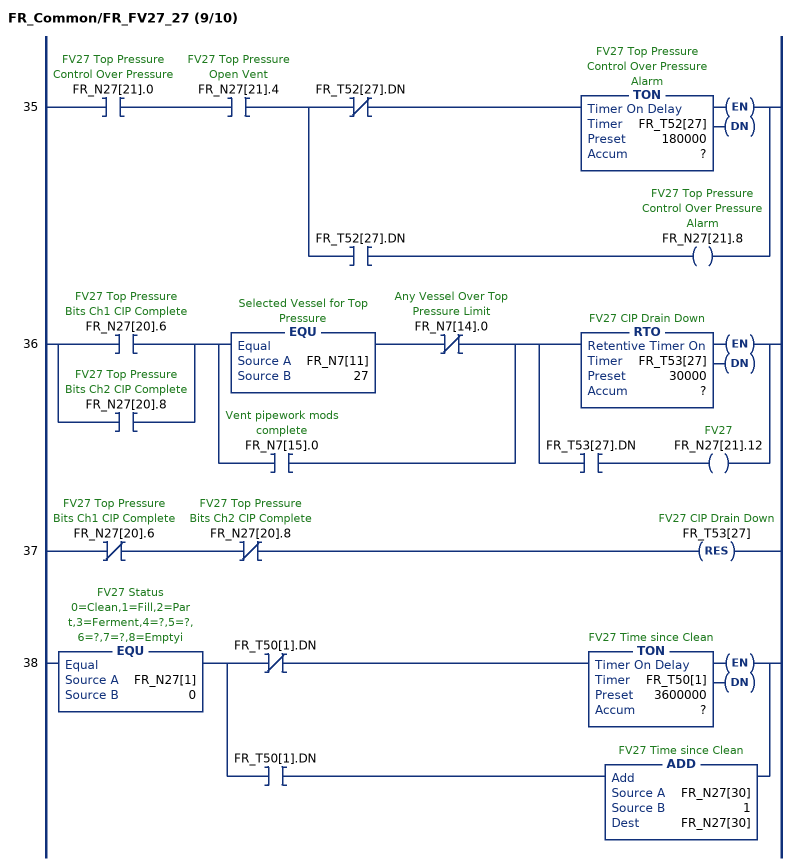
   35: XIC(FR_N27[21].0)XIC(FR_N27[21].4)[XIO(FR_T52[27].DN) TON(FR_T52[27],?,?) ,XIC(FR_T52[27].DN) OTE(FR_N27[21].8) ];
   36: [XIC(FR_N27[20].6) ,XIC(FR_N27[20].8) ][EQU(FR_N7[11],27) XIO(FR_N7[14].0) ,XIC(FR_N7[15].0) ][RTO(FR_T53[27],?,?) ,XIC(FR_T53[27].DN) OTE(FR_N27[21].12) ];
   37: XIO(FR_N27[20].6)XIO(FR_N27[20].8)RES(FR_T53[27]);
   38: EQU(FR_N27[1],0)[XIO(FR_T50[1].DN) TON(FR_T50[1],?,?) ,XIC(FR_T50[1].DN) ADD(FR_N27[30],1,FR_N27[30]) ];
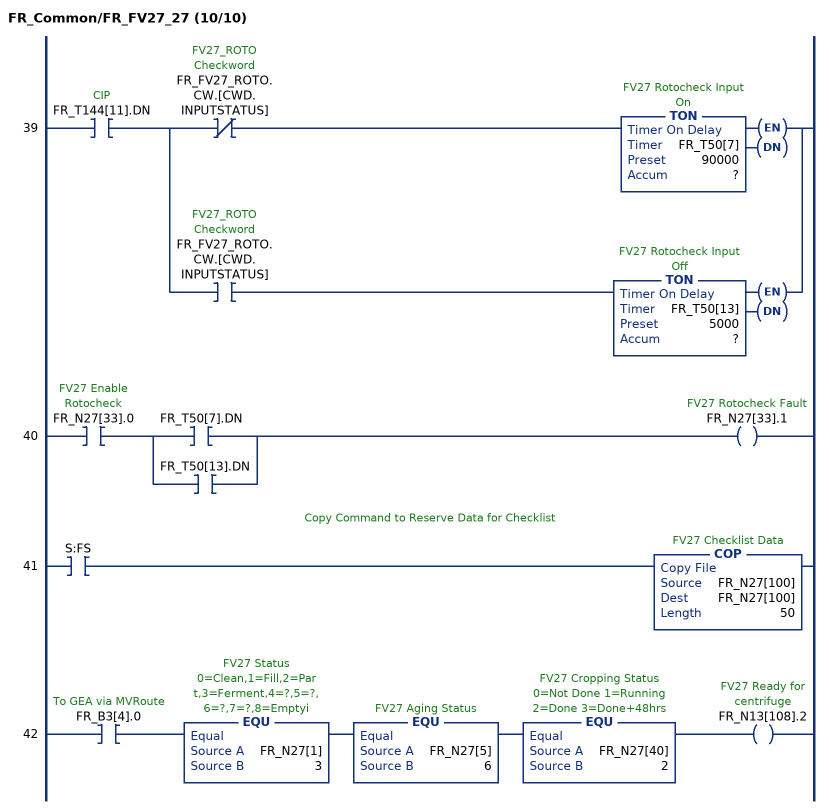
   39: XIC(FR_T144[11].DN)[XIO(FR_FV27_ROTO.CW.[CWD.INPUTSTATUS]) TON(FR_T50[7],?,?) ,XIC(FR_FV27_ROTO.CW.[CWD.INPUTSTATUS]) TON(FR_T50[13],?,?) ];
   40: XIC(FR_N27[33].0)[XIC(FR_T50[7].DN) ,XIC(FR_T50[13].DN) ]OTE(FR_N27[33].1);
   // Copy Command to Reserve Data for Checklist
   41: XIC(S:FS)COP(FR_N27[100],FR_N27[100],50);
   42: XIC(FR_B3[4].0)EQU(FR_N27[1],3)EQU(FR_N27[5],6)EQU(FR_N27[40],2)OTE(FR_N13[108].2);
END_ROUTINE

ROUTINE FR_FV28_28   (* ladder *)
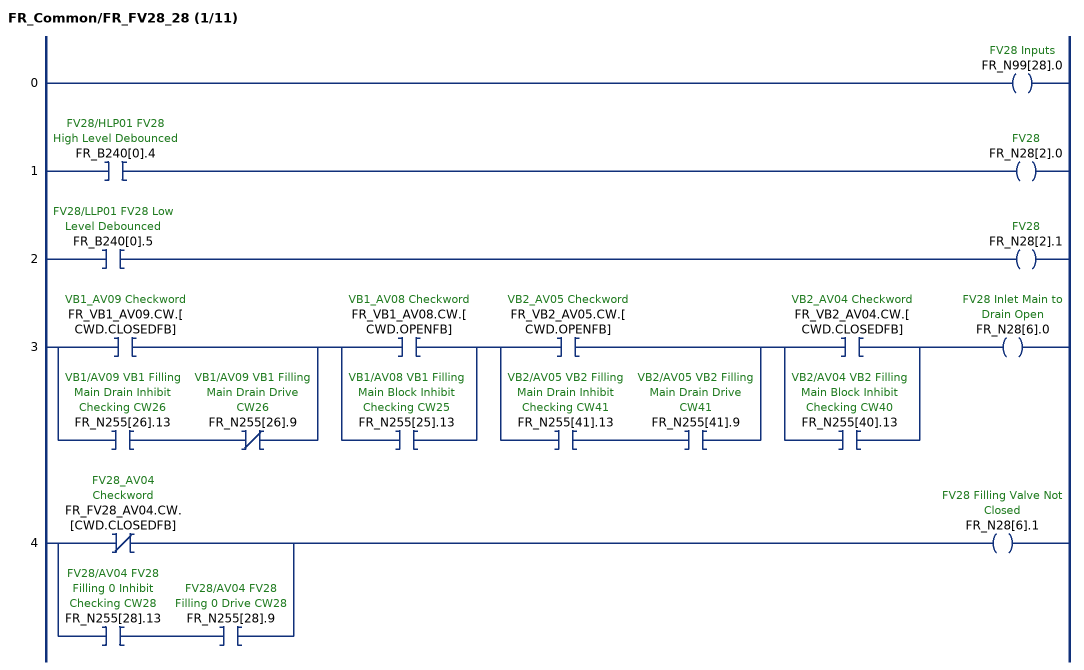
   0: OTE(FR_N99[28].0);
   1: XIC(FR_B240[0].4)OTE(FR_N28[2].0);
   2: XIC(FR_B240[0].5)OTE(FR_N28[2].1);
   3: [XIC(FR_VB1_AV09.CW.[CWD.CLOSEDFB]) ,XIC(FR_N255[26].13) XIO(FR_N255[26].9) ][XIC(FR_VB1_AV08.CW.[CWD.OPENFB]) ,XIC(FR_N255[25].13) ][XIC(FR_VB2_AV05.CW.[CWD.OPENFB]) ,XIC(FR_N255[41].13) XIC(FR_N255[41].9) ][XIC(FR_VB2_AV04.CW.[CWD.CLOSEDFB]) ,XIC(FR_N255[40].13) ]OTE(FR_N28[6].0);
   4: [XIO(FR_FV28_AV04.CW.[CWD.CLOSEDFB]) ,XIC(FR_N255[28].13) XIC(FR_N255[28].9) ]OTE(FR_N28[6].1);
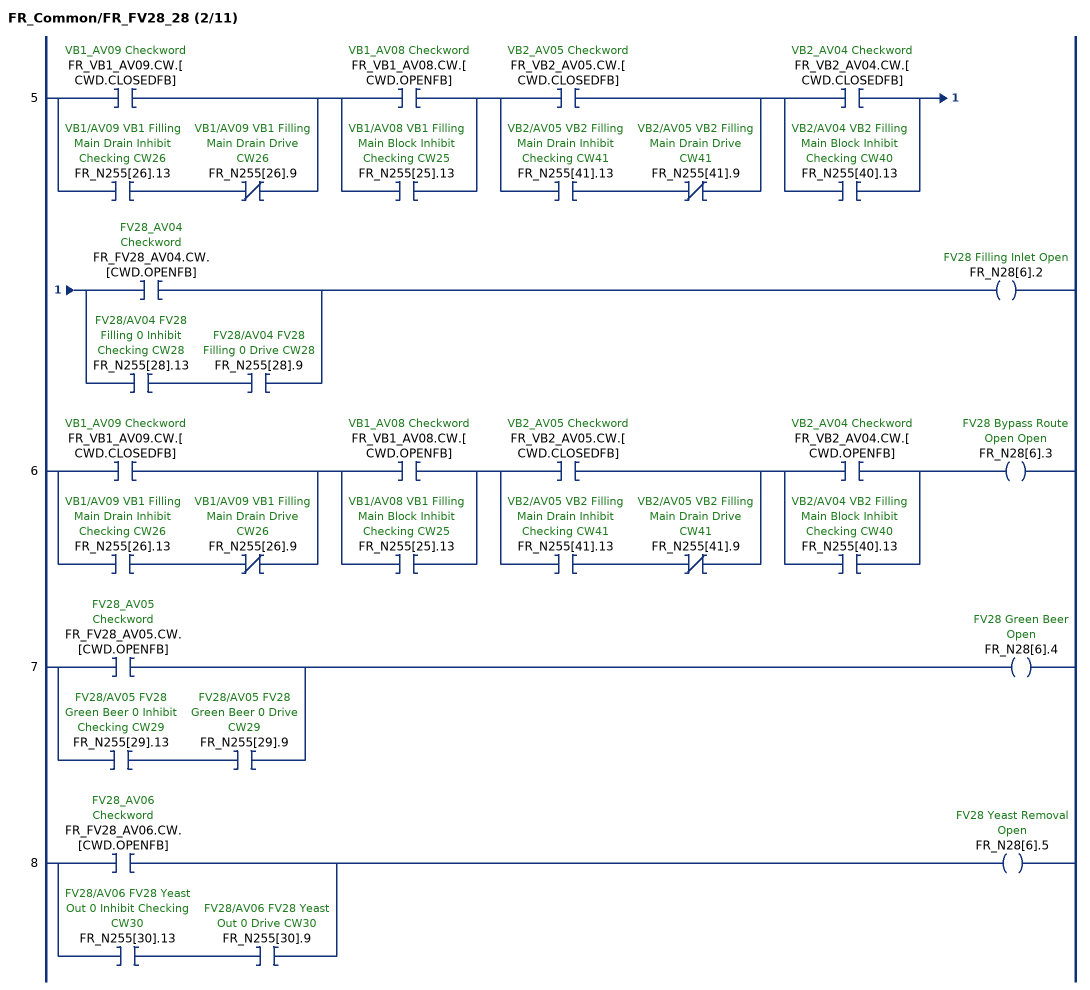
   5: [XIC(FR_VB1_AV09.CW.[CWD.CLOSEDFB]) ,XIC(FR_N255[26].13) XIO(FR_N255[26].9) ][XIC(FR_VB1_AV08.CW.[CWD.OPENFB]) ,XIC(FR_N255[25].13) ][XIC(FR_VB2_AV05.CW.[CWD.CLOSEDFB]) ,XIC(FR_N255[41].13) XIO(FR_N255[41].9) ][XIC(FR_VB2_AV04.CW.[CWD.CLOSEDFB]) ,XIC(FR_N255[40].13) ][XIC(FR_FV28_AV04.CW.[CWD.OPENFB]) ,XIC(FR_N255[28].13) XIC(FR_N255[28].9) ]OTE(FR_N28[6].2);
   6: [XIC(FR_VB1_AV09.CW.[CWD.CLOSEDFB]) ,XIC(FR_N255[26].13) XIO(FR_N255[26].9) ][XIC(FR_VB1_AV08.CW.[CWD.OPENFB]) ,XIC(FR_N255[25].13) ][XIC(FR_VB2_AV05.CW.[CWD.CLOSEDFB]) ,XIC(FR_N255[41].13) XIO(FR_N255[41].9) ][XIC(FR_VB2_AV04.CW.[CWD.OPENFB]) ,XIC(FR_N255[40].13) ]OTE(FR_N28[6].3);
   7: [XIC(FR_FV28_AV05.CW.[CWD.OPENFB]) ,XIC(FR_N255[29].13) XIC(FR_N255[29].9) ]OTE(FR_N28[6].4);
   8: [XIC(FR_FV28_AV06.CW.[CWD.OPENFB]) ,XIC(FR_N255[30].13) XIC(FR_N255[30].9) ]OTE(FR_N28[6].5);
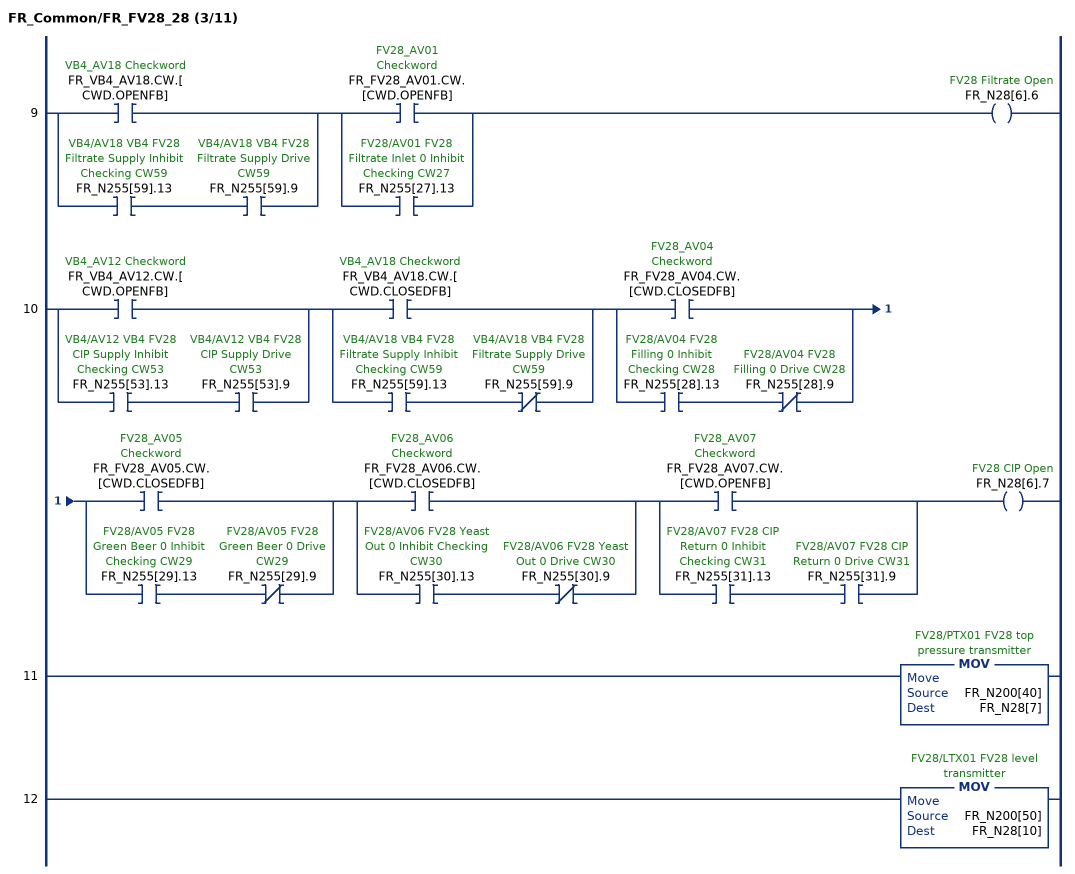
   9: [XIC(FR_VB4_AV18.CW.[CWD.OPENFB]) ,XIC(FR_N255[59].13) XIC(FR_N255[59].9) ][XIC(FR_FV28_AV01.CW.[CWD.OPENFB]) ,XIC(FR_N255[27].13) ]OTE(FR_N28[6].6);
   10: [XIC(FR_VB4_AV12.CW.[CWD.OPENFB]) ,XIC(FR_N255[53].13) XIC(FR_N255[53].9) ][XIC(FR_VB4_AV18.CW.[CWD.CLOSEDFB]) ,XIC(FR_N255[59].13) XIO(FR_N255[59].9) ][XIC(FR_FV28_AV04.CW.[CWD.CLOSEDFB]) ,XIC(FR_N255[28].13) XIO(FR_N255[28].9) ][XIC(FR_FV28_AV05.CW.[CWD.CLOSEDFB]) ,XIC(FR_N255[29].13) XIO(FR_N255[29].9) ][XIC(FR_FV28_AV06.CW.[CWD.CLOSEDFB]) ,XIC(FR_N255[30].13) XIO(FR_N255[30].9) ][XIC(FR_FV28_AV07.CW.[CWD.OPENFB]) ,XIC(FR_N255[31].13) XIC(FR_N255[31].9) ]OTE(FR_N28[6].7);
   11: MOV(FR_N200[40],FR_N28[7]);
   12: MOV(FR_N200[50],FR_N28[10]);
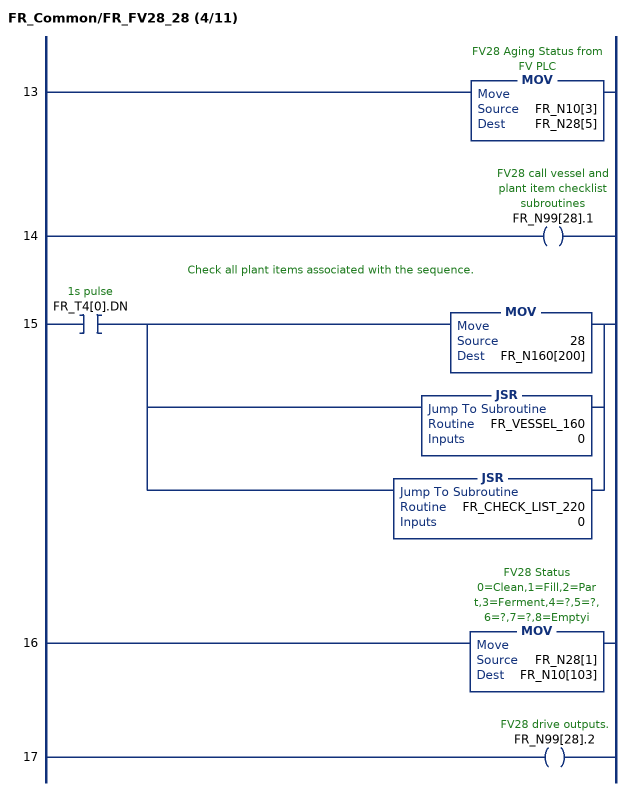
   13: MOV(FR_N10[3],FR_N28[5]);
   14: OTE(FR_N99[28].1);
   // Check all plant items associated with the sequence.
   15: XIC(FR_T4[0].DN)[MOV(28,FR_N160[200]) ,JSR(FR_VESSEL_160,0) ,JSR(FR_CHECK_LIST_220,0) ];
   16: MOV(FR_N28[1],FR_N10[103]);
   17: OTE(FR_N99[28].2);
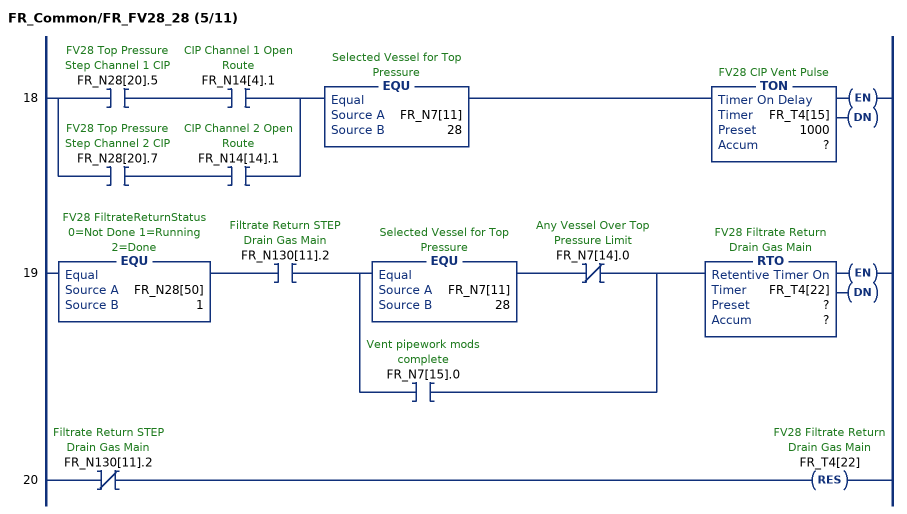
   18: [XIC(FR_N28[20].5) XIC(FR_N14[4].1) ,XIC(FR_N28[20].7) XIC(FR_N14[14].1) ]EQU(FR_N7[11],28)TON(FR_T4[15],?,?);
   19: EQU(FR_N28[50],1)XIC(FR_N130[11].2)[EQU(FR_N7[11],28) XIO(FR_N7[14].0) ,XIC(FR_N7[15].0) ]RTO(FR_T4[22],?,?);
   20: XIO(FR_N130[11].2)RES(FR_T4[22]);
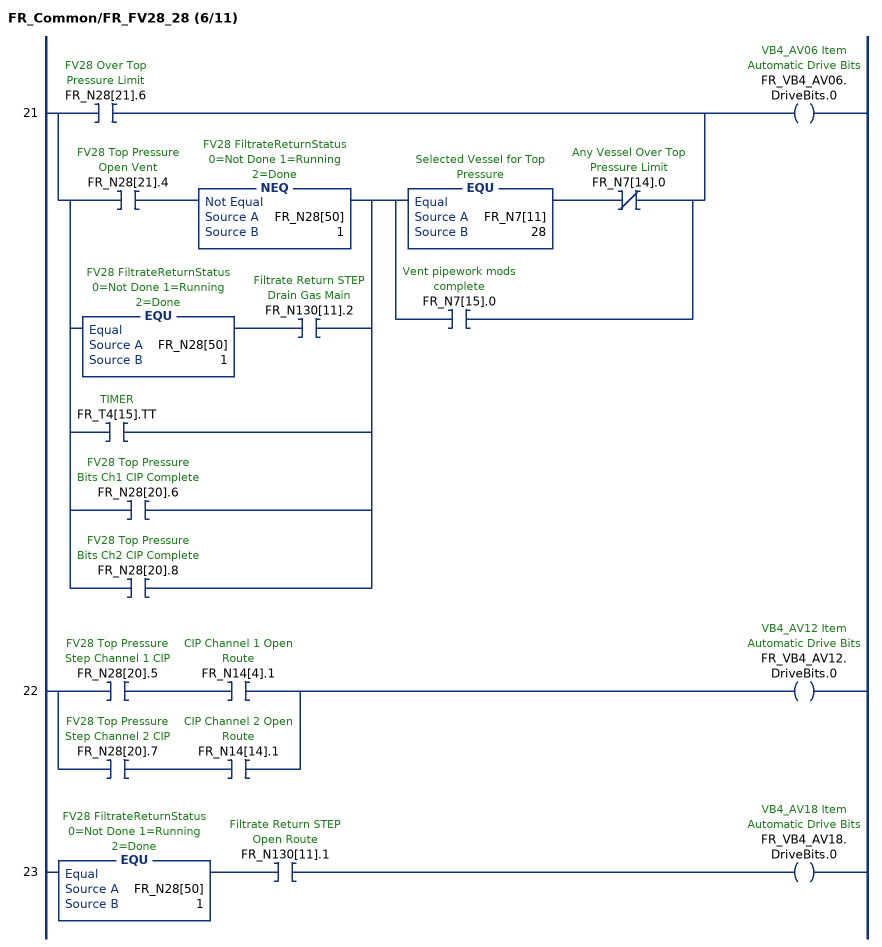
   21: [XIC(FR_N28[21].6) ,[XIC(FR_N28[21].4) NEQ(FR_N28[50],1) ,EQU(FR_N28[50],1) XIC(FR_N130[11].2) ,XIC(FR_T4[15].TT) ,[XIC(FR_N28[20].6) ,XIC(FR_N28[20].8) ] ] [EQU(FR_N7[11],28) XIO(FR_N7[14].0) ,XIC(FR_N7[15].0) ] ]OTE(FR_VB4_AV06.DriveBits.0);
   22: [XIC(FR_N28[20].5) XIC(FR_N14[4].1) ,XIC(FR_N28[20].7) XIC(FR_N14[14].1) ]OTE(FR_VB4_AV12.DriveBits.0);
   23: EQU(FR_N28[50],1)XIC(FR_N130[11].1)OTE(FR_VB4_AV18.DriveBits.0);
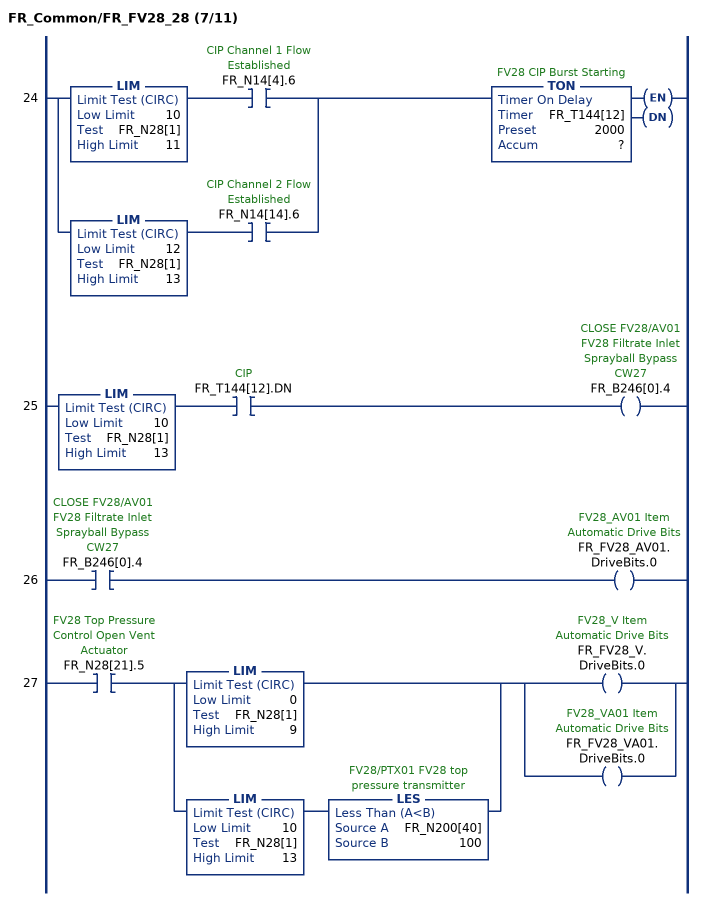
   24: [LIM(10,FR_N28[1],11) XIC(FR_N14[4].6) ,LIM(12,FR_N28[1],13) XIC(FR_N14[14].6) ]TON(FR_T144[12],?,?);
   25: LIM(10,FR_N28[1],13)XIC(FR_T144[12].DN)OTE(FR_B246[0].4);
   26: XIC(FR_B246[0].4)OTE(FR_FV28_AV01.DriveBits.0);
   27: XIC(FR_N28[21].5)[LIM(0,FR_N28[1],9) ,LIM(10,FR_N28[1],13) LES(FR_N200[40],100) ][OTE(FR_FV28_V.DriveBits.0) ,OTE(FR_FV28_VA01.DriveBits.0) ];
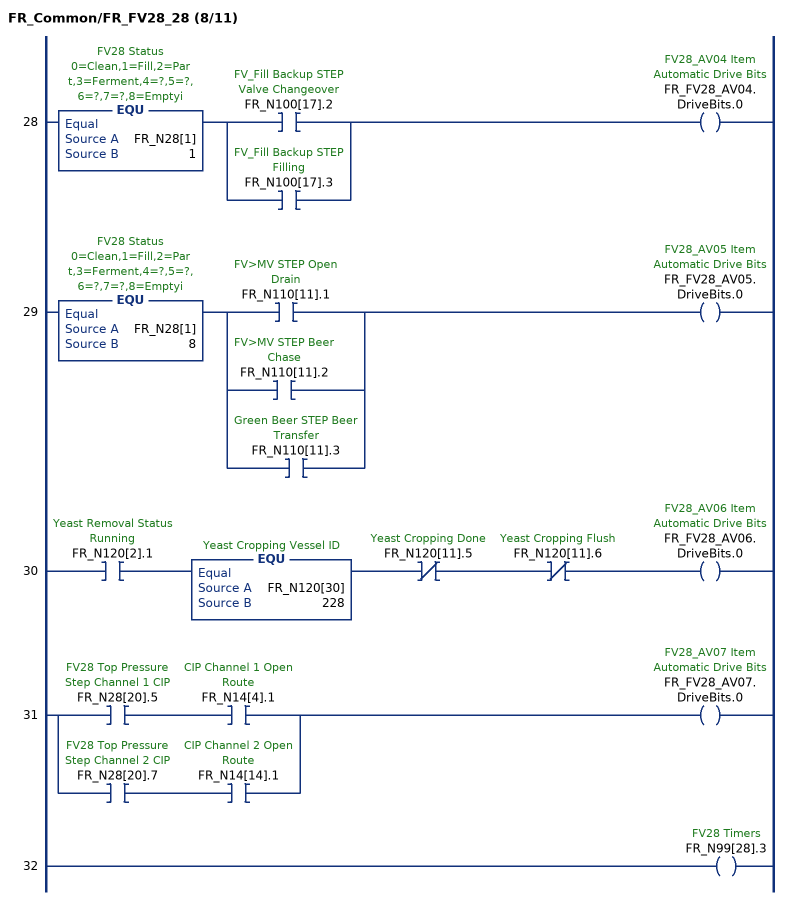
   28: EQU(FR_N28[1],1)[XIC(FR_N100[17].2) ,XIC(FR_N100[17].3) ]OTE(FR_FV28_AV04.DriveBits.0);
   29: EQU(FR_N28[1],8)[XIC(FR_N110[11].1) ,XIC(FR_N110[11].2) ,XIC(FR_N110[11].3) ]OTE(FR_FV28_AV05.DriveBits.0);
   30: XIC(FR_N120[2].1)EQU(FR_N120[30],228)XIO(FR_N120[11].5)XIO(FR_N120[11].6)OTE(FR_FV28_AV06.DriveBits.0);
   31: [XIC(FR_N28[20].5) XIC(FR_N14[4].1) ,XIC(FR_N28[20].7) XIC(FR_N14[14].1) ]OTE(FR_FV28_AV07.DriveBits.0);
   32: OTE(FR_N99[28].3);
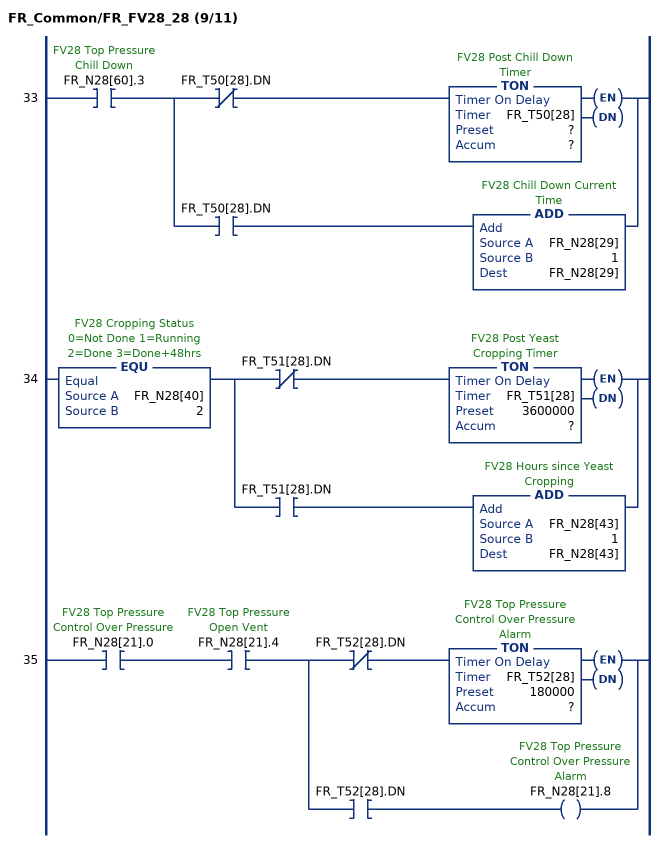
   33: XIC(FR_N28[60].3)[XIO(FR_T50[28].DN) TON(FR_T50[28],?,?) ,XIC(FR_T50[28].DN) ADD(FR_N28[29],1,FR_N28[29]) ];
   34: EQU(FR_N28[40],2)[XIO(FR_T51[28].DN) TON(FR_T51[28],?,?) ,XIC(FR_T51[28].DN) ADD(FR_N28[43],1,FR_N28[43]) ];
   35: XIC(FR_N28[21].0)XIC(FR_N28[21].4)[XIO(FR_T52[28].DN) TON(FR_T52[28],?,?) ,XIC(FR_T52[28].DN) OTE(FR_N28[21].8) ];
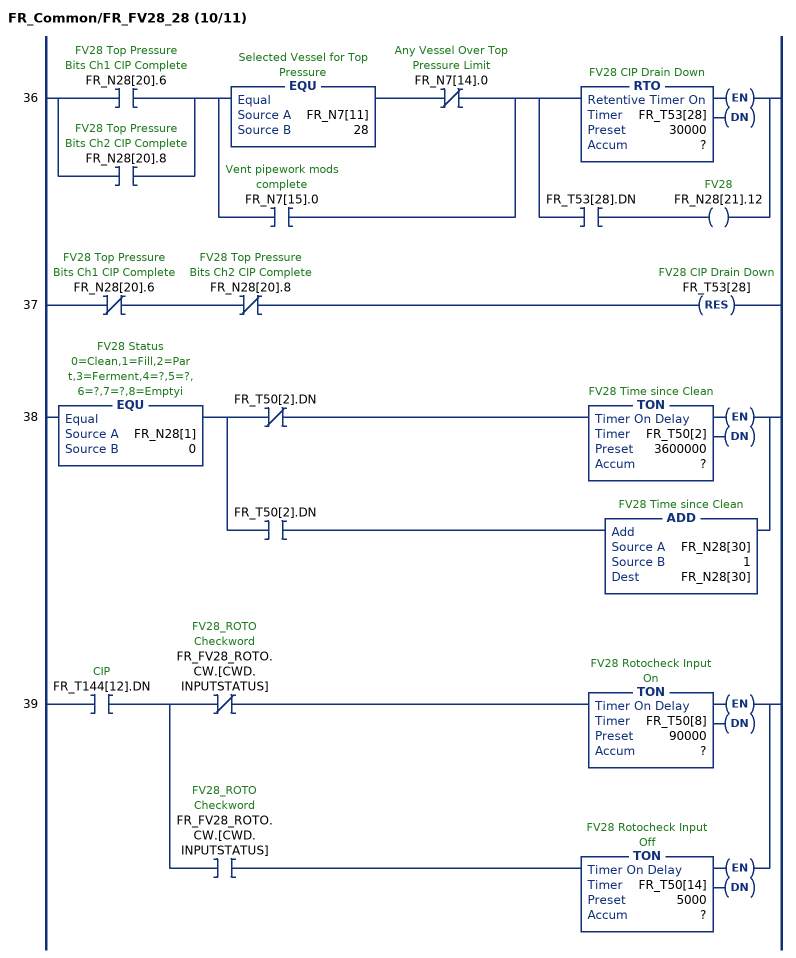
   36: [XIC(FR_N28[20].6) ,XIC(FR_N28[20].8) ][EQU(FR_N7[11],28) XIO(FR_N7[14].0) ,XIC(FR_N7[15].0) ][RTO(FR_T53[28],?,?) ,XIC(FR_T53[28].DN) OTE(FR_N28[21].12) ];
   37: XIO(FR_N28[20].6)XIO(FR_N28[20].8)RES(FR_T53[28]);
   38: EQU(FR_N28[1],0)[XIO(FR_T50[2].DN) TON(FR_T50[2],?,?) ,XIC(FR_T50[2].DN) ADD(FR_N28[30],1,FR_N28[30]) ];
   39: XIC(FR_T144[12].DN)[XIO(FR_FV28_ROTO.CW.[CWD.INPUTSTATUS]) TON(FR_T50[8],?,?) ,XIC(FR_FV28_ROTO.CW.[CWD.INPUTSTATUS]) TON(FR_T50[14],?,?) ];
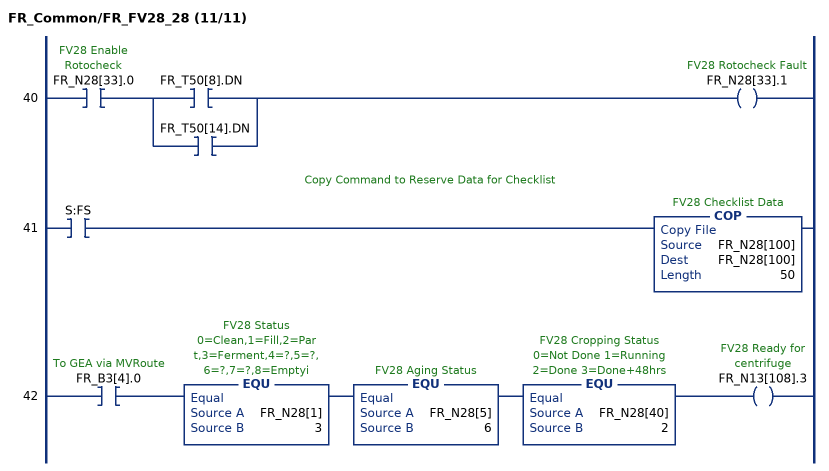
   40: XIC(FR_N28[33].0)[XIC(FR_T50[8].DN) ,XIC(FR_T50[14].DN) ]OTE(FR_N28[33].1);
   // Copy Command to Reserve Data for Checklist
   41: XIC(S:FS)COP(FR_N28[100],FR_N28[100],50);
   42: XIC(FR_B3[4].0)EQU(FR_N28[1],3)EQU(FR_N28[5],6)EQU(FR_N28[40],2)OTE(FR_N13[108].3);
END_ROUTINE
